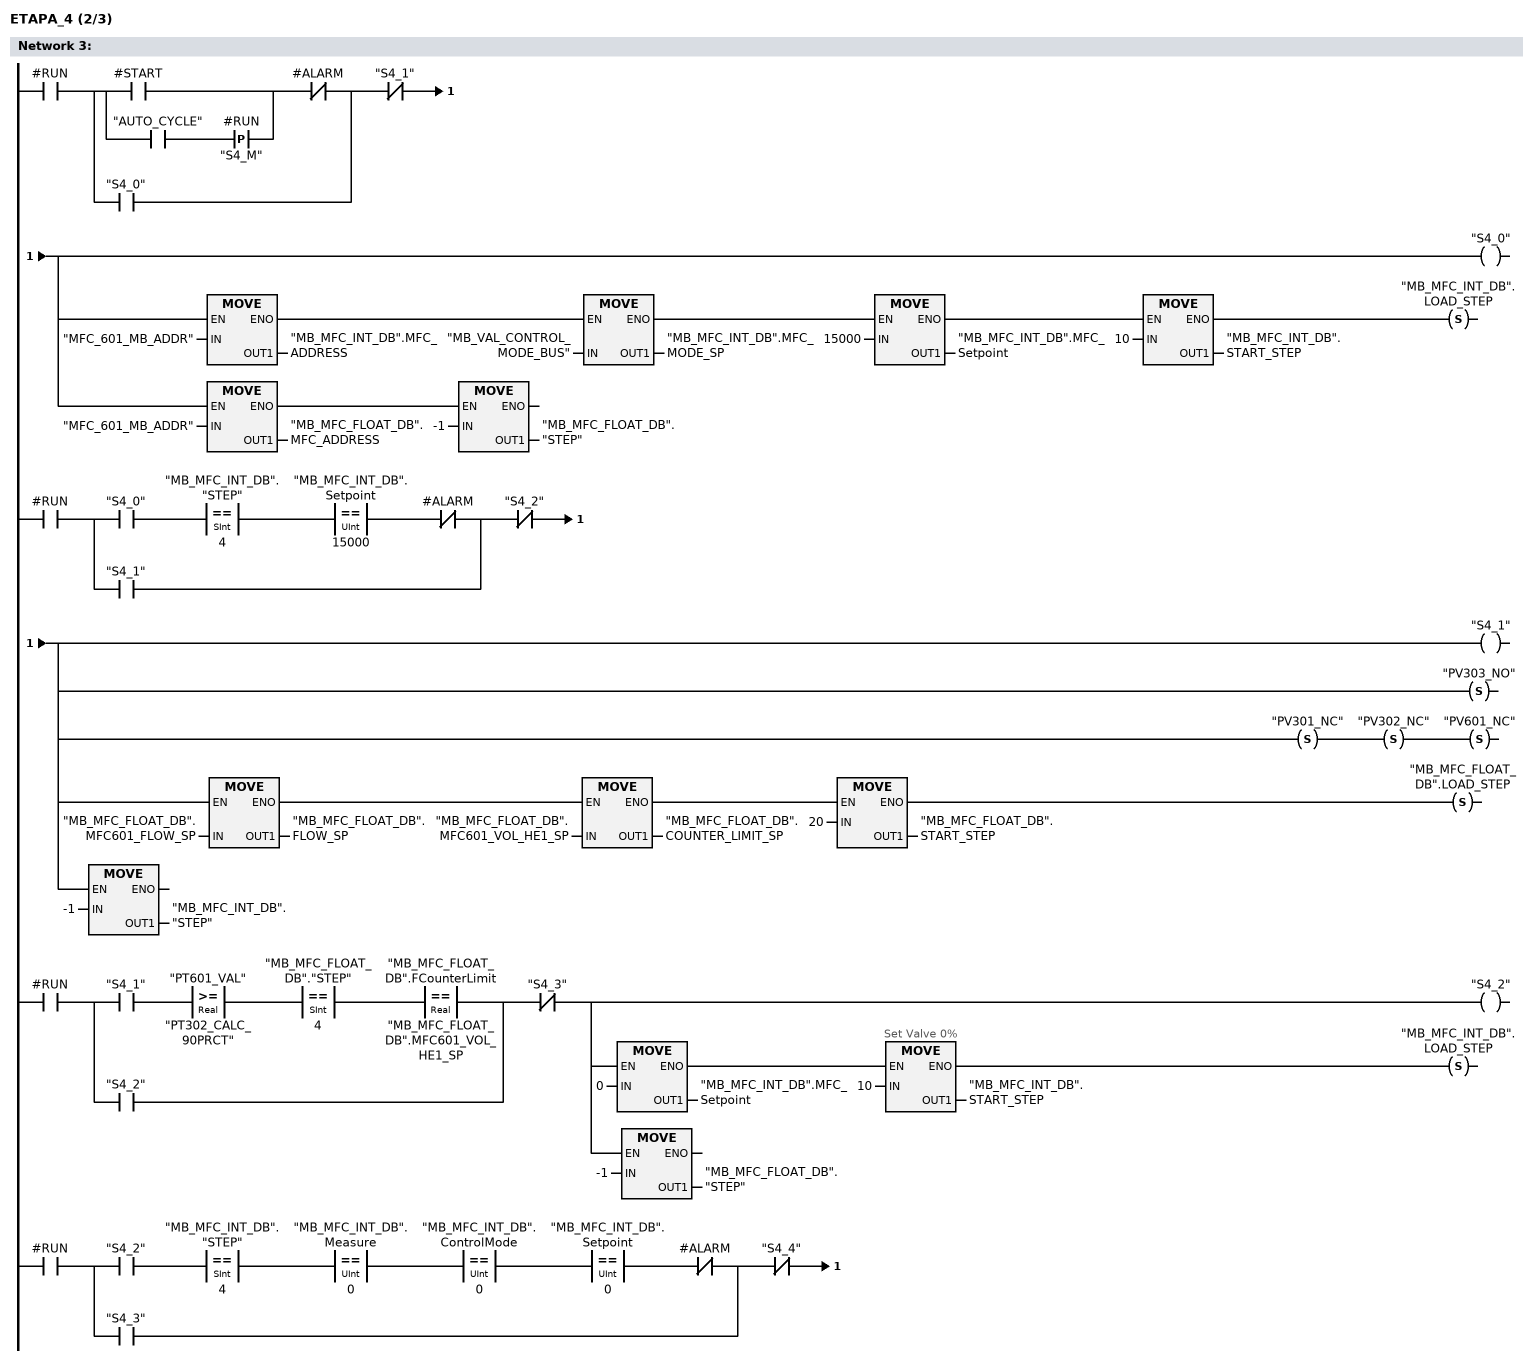
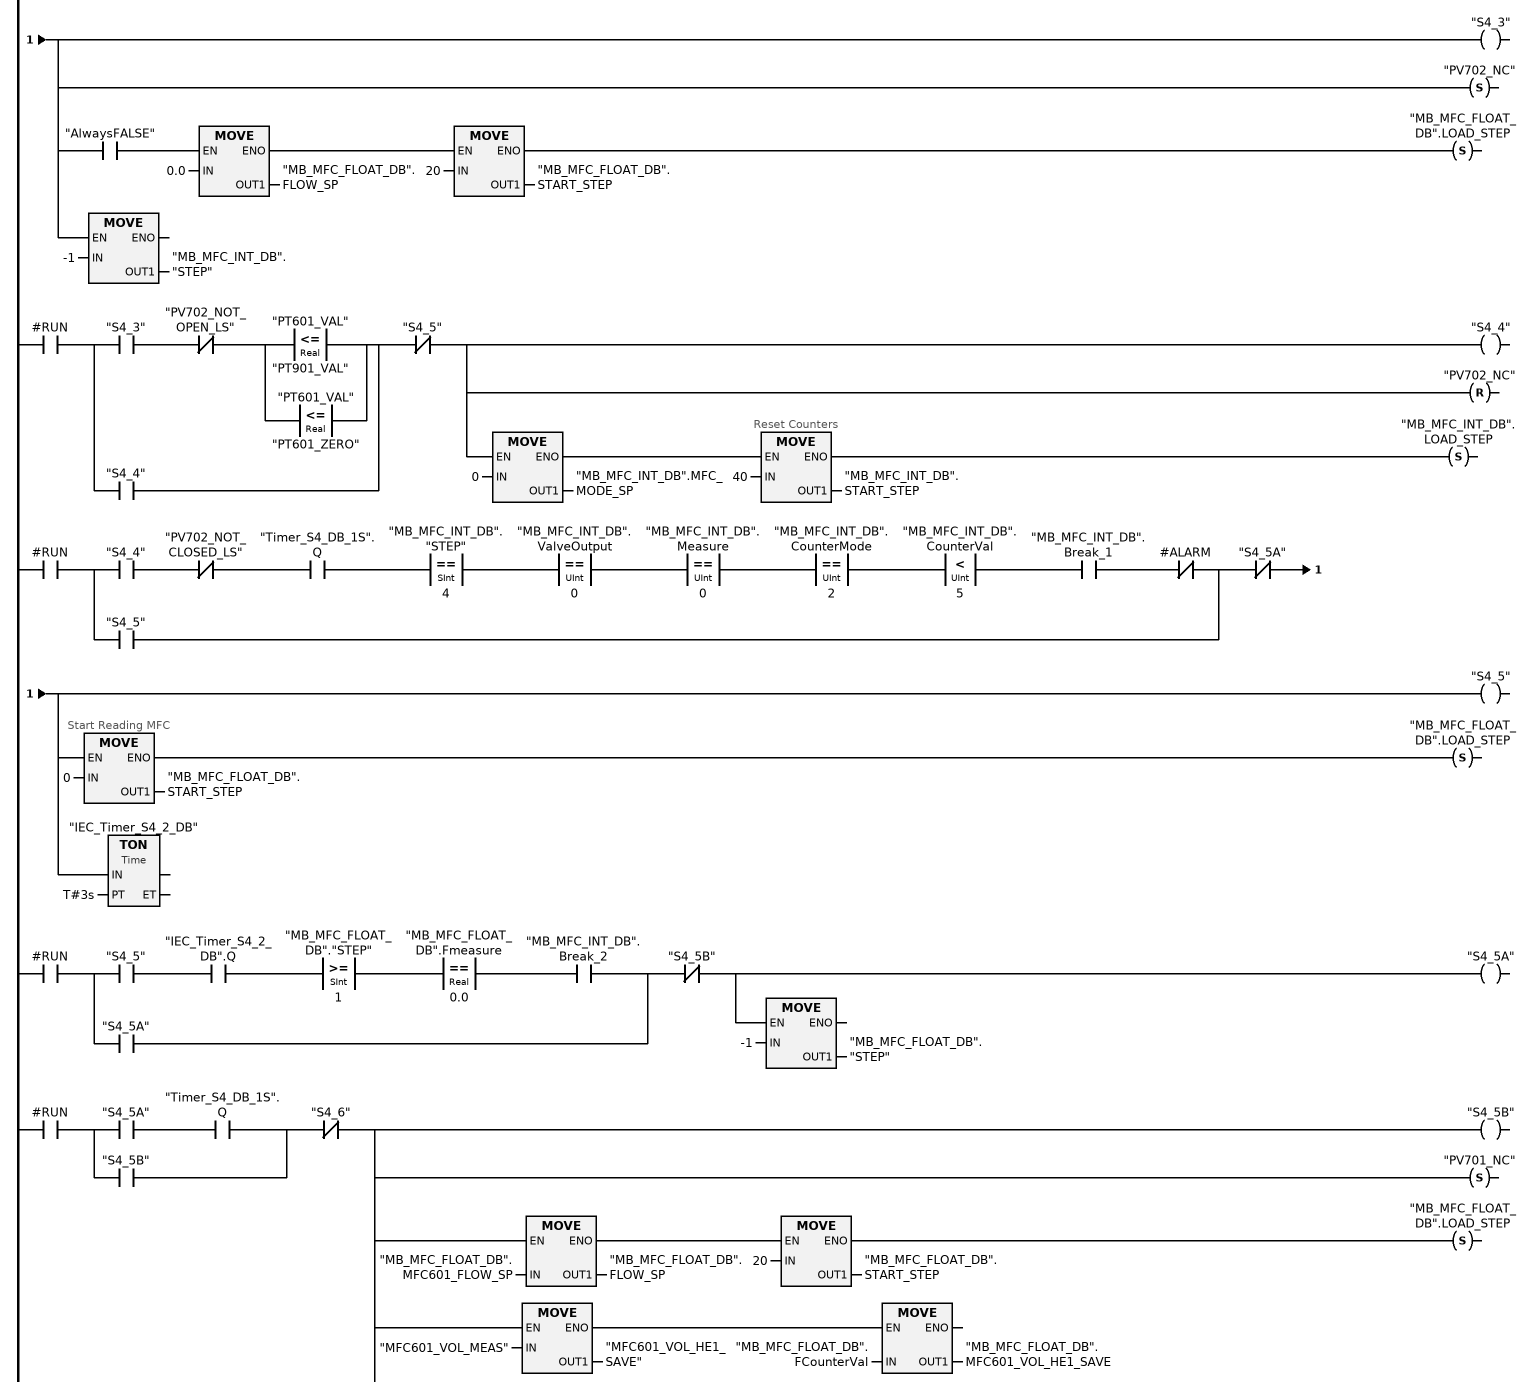
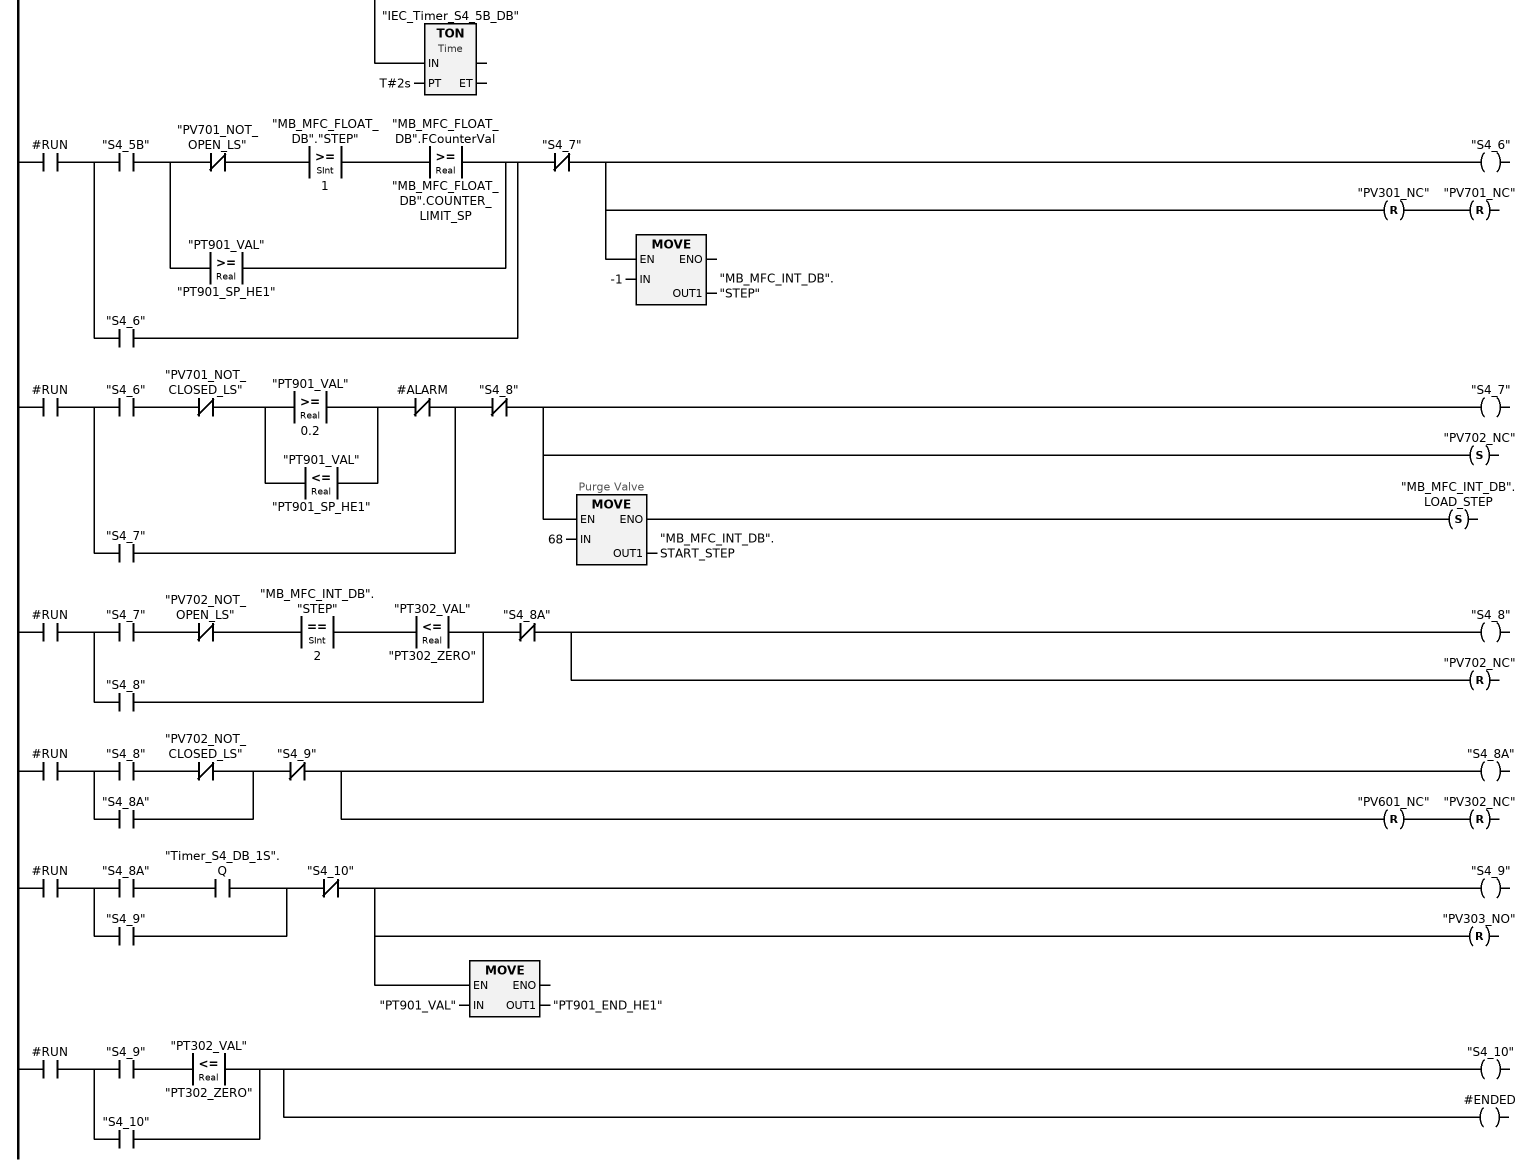
   #_w1 := #RUN AND "AUTO_CYCLE" AND #RUN AND NOT "S4_M";   // rising edge of #RUN
   "S4_M" := #RUN;
   "S4_0" := ((((#RUN AND #START) OR #_w1) AND NOT #ALARM) OR (#RUN AND "S4_0")) AND NOT "S4_1";
   IF "S4_0" THEN
       "MB_MFC_INT_DB".MFC_ADDRESS := "MFC_601_MB_ADDR";
       "MB_MFC_INT_DB".MFC_MODE_SP := "MB_VAL_CONTROL_MODE_BUS";
       "MB_MFC_INT_DB".MFC_Setpoint := 15000;
       "MB_MFC_INT_DB".START_STEP := 10;
       "MB_MFC_INT_DB".LOAD_STEP := TRUE;
       "MB_MFC_FLOAT_DB".MFC_ADDRESS := "MFC_601_MB_ADDR";
       "MB_MFC_FLOAT_DB"."STEP" := -1;
   END_IF;
   "S4_1" := #RUN AND (("S4_0" AND ("MB_MFC_INT_DB"."STEP" = 4) AND ("MB_MFC_INT_DB".Setpoint = 15000) AND NOT #ALARM) OR "S4_1") AND NOT "S4_2";
   IF "S4_1" THEN
       "PV303_NO" := TRUE;
       "PV301_NC" := TRUE;
       "PV302_NC" := TRUE;
       "PV601_NC" := TRUE;
       "MB_MFC_FLOAT_DB".FLOW_SP := "MB_MFC_FLOAT_DB".MFC601_FLOW_SP;
       "MB_MFC_FLOAT_DB".COUNTER_LIMIT_SP := "MB_MFC_FLOAT_DB".MFC601_VOL_HE1_SP;
       "MB_MFC_FLOAT_DB".START_STEP := 20;
       "MB_MFC_FLOAT_DB".LOAD_STEP := TRUE;
       "MB_MFC_INT_DB"."STEP" := -1;
   END_IF;
   "S4_2" := #RUN AND (("S4_1" AND ("PT601_VAL" >= "PT302_CALC_90PRCT") AND ("MB_MFC_FLOAT_DB"."STEP" = 4) AND ("MB_MFC_FLOAT_DB".FCounterLimit = "MB_MFC_FLOAT_DB".MFC601_VOL_HE1_SP)) OR "S4_2") AND NOT "S4_3";
   IF "S4_2" THEN
       "MB_MFC_INT_DB".MFC_Setpoint := 0;
       "MB_MFC_INT_DB".START_STEP := 10;   // Set Valve 0%
       "MB_MFC_INT_DB".LOAD_STEP := TRUE;
       "MB_MFC_FLOAT_DB"."STEP" := -1;
   END_IF;
   "S4_3" := #RUN AND (("S4_2" AND ("MB_MFC_INT_DB"."STEP" = 4) AND ("MB_MFC_INT_DB".Measure = 0) AND ("MB_MFC_INT_DB".ControlMode = 0) AND ("MB_MFC_INT_DB".Setpoint = 0) AND NOT #ALARM) OR "S4_3") AND NOT "S4_4";
   IF "S4_3" THEN "PV702_NC" := TRUE; END_IF;
   IF "S4_3" AND "AlwaysFALSE" THEN
       "MB_MFC_FLOAT_DB".FLOW_SP := 0.0;
       "MB_MFC_FLOAT_DB".START_STEP := 20;
       "MB_MFC_FLOAT_DB".LOAD_STEP := TRUE;
   END_IF;
   IF "S4_3" THEN "MB_MFC_INT_DB"."STEP" := -1; END_IF;
   "S4_4" := #RUN AND (("S4_3" AND NOT "PV702_NOT_OPEN_LS" AND (("PT601_VAL" <= "PT901_VAL") OR ("PT601_VAL" <= "PT601_ZERO"))) OR "S4_4") AND NOT "S4_5";
   IF "S4_4" THEN
       "PV702_NC" := FALSE;
       "MB_MFC_INT_DB".MFC_MODE_SP := 0;
       "MB_MFC_INT_DB".START_STEP := 40;   // Reset Counters
       "MB_MFC_INT_DB".LOAD_STEP := TRUE;
   END_IF;
   "S4_5" := #RUN AND (("S4_4" AND NOT "PV702_NOT_CLOSED_LS" AND "Timer_S4_DB_1S".Q AND ("MB_MFC_INT_DB"."STEP" = 4) AND ("MB_MFC_INT_DB".ValveOutput = 0) AND ("MB_MFC_INT_DB".Measure = 0) AND ("MB_MFC_INT_DB".CounterMode = 2) AND ("MB_MFC_INT_DB".CounterVal < 5) AND "MB_MFC_INT_DB".Break_1 AND NOT #ALARM) OR "S4_5") AND NOT "S4_5A";
   IF "S4_5" THEN
       "MB_MFC_FLOAT_DB".START_STEP := 0;   // Start Reading MFC
       "MB_MFC_FLOAT_DB".LOAD_STEP := TRUE;
   END_IF;
   "IEC_Timer_S4_2_DB".TON(IN := "S4_5", PT := T#3s);
   "S4_5A" := #RUN AND (("S4_5" AND "IEC_Timer_S4_2_DB".Q AND ("MB_MFC_FLOAT_DB"."STEP" >= 1) AND ("MB_MFC_FLOAT_DB".Fmeasure = 0.0) AND "MB_MFC_INT_DB".Break_2) OR "S4_5A") AND NOT "S4_5B";
   IF "S4_5A" THEN "MB_MFC_FLOAT_DB"."STEP" := -1; END_IF;
   "S4_5B" := #RUN AND (("S4_5A" AND "Timer_S4_DB_1S".Q) OR "S4_5B") AND NOT "S4_6";
   IF "S4_5B" THEN
       "PV701_NC" := TRUE;
       "MB_MFC_FLOAT_DB".FLOW_SP := "MB_MFC_FLOAT_DB".MFC601_FLOW_SP;
       "MB_MFC_FLOAT_DB".START_STEP := 20;
       "MB_MFC_FLOAT_DB".LOAD_STEP := TRUE;
       "MFC601_VOL_HE1_SAVE" := "MFC601_VOL_MEAS";
       "MB_MFC_FLOAT_DB".MFC601_VOL_HE1_SAVE := "MB_MFC_FLOAT_DB".FCounterVal;
   END_IF;
   "IEC_Timer_S4_5B_DB".TON(IN := "S4_5B", PT := T#2s);
   "S4_6" := #RUN AND (("S4_5B" AND ((NOT "PV701_NOT_OPEN_LS" AND ("MB_MFC_FLOAT_DB"."STEP" >= 1) AND ("MB_MFC_FLOAT_DB".FCounterVal >= "MB_MFC_FLOAT_DB".COUNTER_LIMIT_SP)) OR ("PT901_VAL" >= "PT901_SP_HE1"))) OR "S4_6") AND NOT "S4_7";
   IF "S4_6" THEN
       "PV301_NC" := FALSE;
       "PV701_NC" := FALSE;
       "MB_MFC_INT_DB"."STEP" := -1;
   END_IF;
   "S4_7" := #RUN AND (("S4_6" AND NOT "PV701_NOT_CLOSED_LS" AND (("PT901_VAL" >= 0.2) OR ("PT901_VAL" <= "PT901_SP_HE1")) AND NOT #ALARM) OR "S4_7") AND NOT "S4_8";
   IF "S4_7" THEN
       "PV702_NC" := TRUE;
       "MB_MFC_INT_DB".START_STEP := 68;   // Purge Valve
       "MB_MFC_INT_DB".LOAD_STEP := TRUE;
   END_IF;
   "S4_8" := #RUN AND (("S4_7" AND NOT "PV702_NOT_OPEN_LS" AND ("MB_MFC_INT_DB"."STEP" = 2) AND ("PT302_VAL" <= "PT302_ZERO")) OR "S4_8") AND NOT "S4_8A";
   IF "S4_8" THEN "PV702_NC" := FALSE; END_IF;
   "S4_8A" := #RUN AND (("S4_8" AND NOT "PV702_NOT_CLOSED_LS") OR "S4_8A") AND NOT "S4_9";
   IF "S4_8A" THEN
       "PV601_NC" := FALSE;
       "PV302_NC" := FALSE;
   END_IF;
   "S4_9" := #RUN AND (("S4_8A" AND "Timer_S4_DB_1S".Q) OR "S4_9") AND NOT "S4_10";
   IF "S4_9" THEN
       "PV303_NO" := FALSE;
       "PT901_END_HE1" := "PT901_VAL";
   END_IF;
   "S4_10" := #RUN AND (("S4_9" AND ("PT302_VAL" <= "PT302_ZERO")) OR "S4_10");
   #ENDED := "S4_10";
END_REGION

REGION Network 4
   // Timers
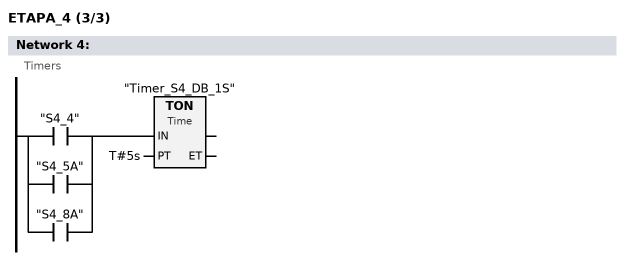
   "Timer_S4_DB_1S".TON(IN := "S4_4" OR "S4_5A" OR "S4_8A", PT := T#5s);
END_REGION
END_FUNCTION

FUNCTION "ETAPA_5" : Void   // FC6, LAD
{ S7_Optimized_Access := 'FALSE' }
VERSION : 0.1
// CICLO de INJECÇÃO - Varrimento Helio 2
   VAR_TEMP   // added for the SCL form of the ladder/FBD networks
      _w1 : Bool;
   END_VAR
BEGIN

REGION Network 1
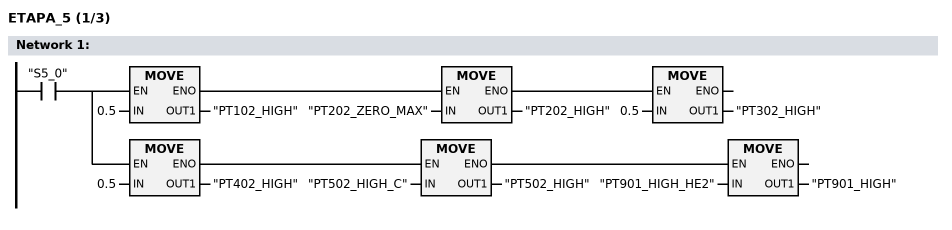
   RUNG wire#powerrail
      Contact( "S5_0" )
      wire#w1
      { S7_GenerateENO := "TRUE" } Move(in := 0.5, out1 => "PT102_HIGH")
      { S7_GenerateENO := "TRUE" } Move(in := "PT202_ZERO_MAX", out1 => "PT202_HIGH")
      { S7_GenerateENO := "TRUE" } Move(in := 0.5, out1 => "PT302_HIGH")
   END_RUNG
   RUNG wire#w1
      { S7_GenerateENO := "TRUE" } Move(in := 0.5, out1 => "PT402_HIGH")
      { S7_GenerateENO := "TRUE" } Move(in := "PT502_HIGH_C", out1 => "PT502_HIGH")
      { S7_GenerateENO := "TRUE" } Move(in := "PT901_HIGH_HE2", out1 => "PT901_HIGH")
   END_RUNG
   // the same network as SCL:
   // ENO of a box is taken as its EN; it also drops when the box reports an error
   IF "S5_0" THEN
       "PT102_HIGH" := 0.5;
       "PT202_HIGH" := "PT202_ZERO_MAX";
       "PT302_HIGH" := 0.5;
       "PT402_HIGH" := 0.5;
       "PT502_HIGH" := "PT502_HIGH_C";
       "PT901_HIGH" := "PT901_HIGH_HE2";
   END_IF;
END_REGION

REGION Network 2
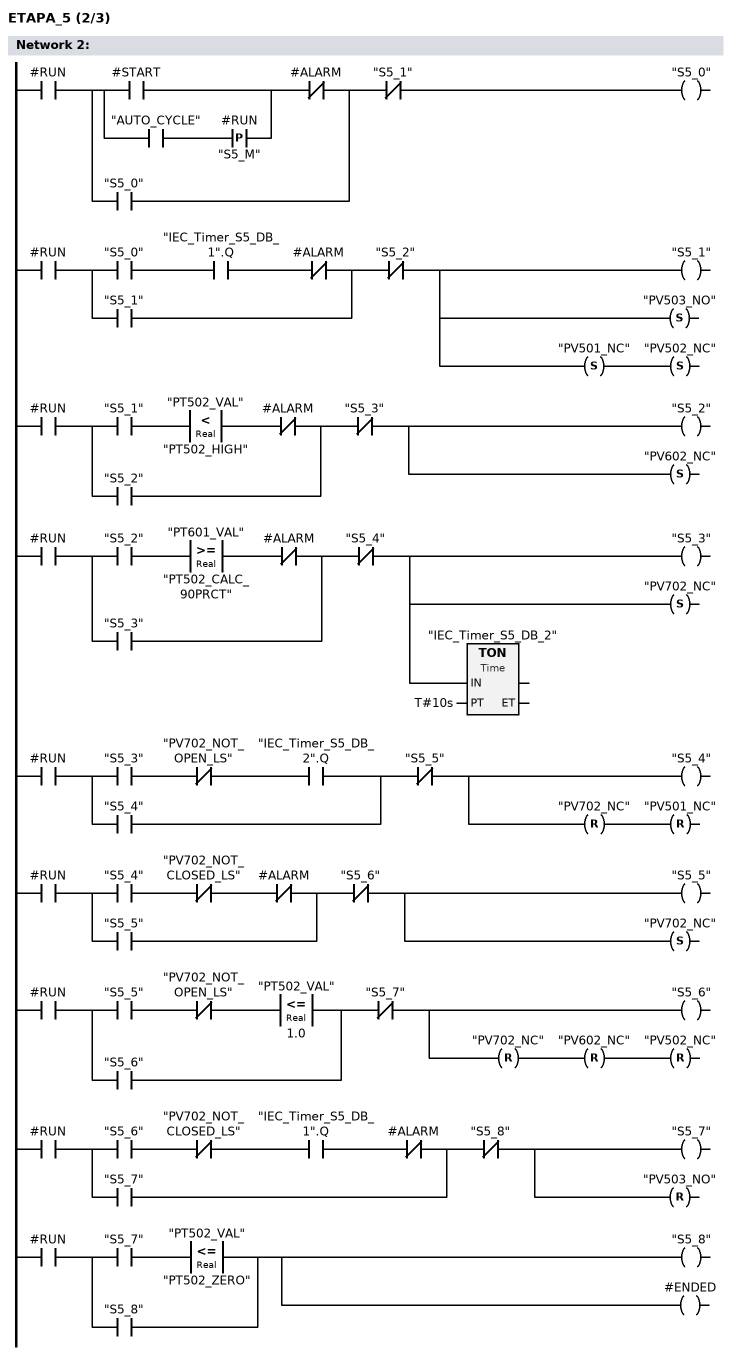
   #_w1 := #RUN AND "AUTO_CYCLE" AND #RUN AND NOT "S5_M";   // rising edge of #RUN
   "S5_M" := #RUN;
   "S5_0" := ((((#RUN AND #START) OR #_w1) AND NOT #ALARM) OR (#RUN AND "S5_0")) AND NOT "S5_1";
   "S5_1" := #RUN AND (("S5_0" AND "IEC_Timer_S5_DB_1".Q AND NOT #ALARM) OR "S5_1") AND NOT "S5_2";
   IF "S5_1" THEN
       "PV503_NO" := TRUE;
       "PV501_NC" := TRUE;
       "PV502_NC" := TRUE;
   END_IF;
   "S5_2" := #RUN AND (("S5_1" AND ("PT502_VAL" < "PT502_HIGH") AND NOT #ALARM) OR "S5_2") AND NOT "S5_3";
   IF "S5_2" THEN "PV602_NC" := TRUE; END_IF;
   "S5_3" := #RUN AND (("S5_2" AND ("PT601_VAL" >= "PT502_CALC_90PRCT") AND NOT #ALARM) OR "S5_3") AND NOT "S5_4";
   IF "S5_3" THEN "PV702_NC" := TRUE; END_IF;
   "IEC_Timer_S5_DB_2".TON(IN := "S5_3", PT := T#10s);
   "S5_4" := #RUN AND (("S5_3" AND NOT "PV702_NOT_OPEN_LS" AND "IEC_Timer_S5_DB_2".Q) OR "S5_4") AND NOT "S5_5";
   IF "S5_4" THEN
       "PV702_NC" := FALSE;
       "PV501_NC" := FALSE;
   END_IF;
   "S5_5" := #RUN AND (("S5_4" AND NOT "PV702_NOT_CLOSED_LS" AND NOT #ALARM) OR "S5_5") AND NOT "S5_6";
   IF "S5_5" THEN "PV702_NC" := TRUE; END_IF;
   "S5_6" := #RUN AND (("S5_5" AND NOT "PV702_NOT_OPEN_LS" AND ("PT502_VAL" <= 1.0)) OR "S5_6") AND NOT "S5_7";
   IF "S5_6" THEN
       "PV702_NC" := FALSE;
       "PV602_NC" := FALSE;
       "PV502_NC" := FALSE;
   END_IF;
   "S5_7" := #RUN AND (("S5_6" AND NOT "PV702_NOT_CLOSED_LS" AND "IEC_Timer_S5_DB_1".Q AND NOT #ALARM) OR "S5_7") AND NOT "S5_8";
   IF "S5_7" THEN "PV503_NO" := FALSE; END_IF;
   "S5_8" := #RUN AND (("S5_7" AND ("PT502_VAL" <= "PT502_ZERO")) OR "S5_8");
   #ENDED := "S5_8";
END_REGION

REGION Network 3
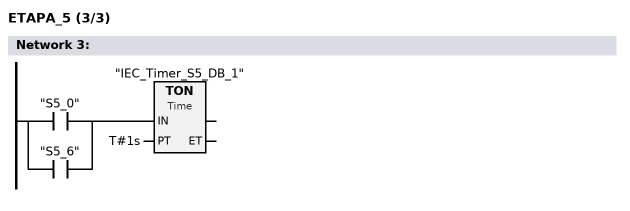
   "IEC_Timer_S5_DB_1".TON(IN := "S5_0" OR "S5_6", PT := T#1s);
END_REGION
END_FUNCTION

FUNCTION "ETAPA_6" : Void   // FC7, LAD
{ S7_Optimized_Access := 'FALSE' }
VERSION : 0.1
// CICLO de INJECÇÃO - injecção de Hidrogénio
   VAR_TEMP   // added for the SCL form of the ladder/FBD networks
      _w1 : Bool;
   END_VAR
BEGIN

REGION Network 1
   // Alarm PT Set Points
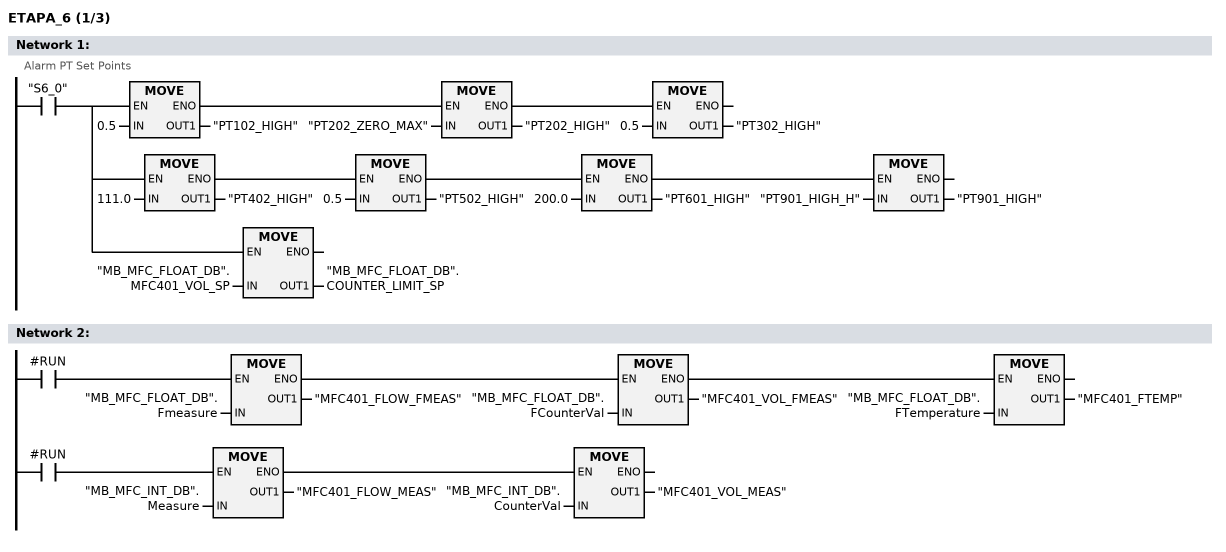
   RUNG wire#powerrail
      Contact( "S6_0" )
      wire#w1
      { S7_GenerateENO := "TRUE" } Move(in := 0.5, out1 => "PT102_HIGH")
      { S7_GenerateENO := "TRUE" } Move(in := "PT202_ZERO_MAX", out1 => "PT202_HIGH")
      { S7_GenerateENO := "TRUE" } Move(in := 0.5, out1 => "PT302_HIGH")
   END_RUNG
   RUNG wire#w1
      { S7_GenerateENO := "TRUE" } Move(in := 111.0, out1 => "PT402_HIGH")
      { S7_GenerateENO := "TRUE" } Move(in := 0.5, out1 => "PT502_HIGH")
      { S7_GenerateENO := "TRUE" } Move(in := 200.0, out1 => "PT601_HIGH")
      { S7_GenerateENO := "TRUE" } Move(in := "PT901_HIGH_H", out1 => "PT901_HIGH")
   END_RUNG
   RUNG wire#w1
      Move(in := "MB_MFC_FLOAT_DB".MFC401_VOL_SP, out1 => "MB_MFC_FLOAT_DB".COUNTER_LIMIT_SP)
   END_RUNG
   // the same network as SCL:
   // ENO of a box is taken as its EN; it also drops when the box reports an error
   IF "S6_0" THEN
       "PT102_HIGH" := 0.5;
       "PT202_HIGH" := "PT202_ZERO_MAX";
       "PT302_HIGH" := 0.5;
       "PT402_HIGH" := 111.0;
       "PT502_HIGH" := 0.5;
       "PT601_HIGH" := 200.0;
       "PT901_HIGH" := "PT901_HIGH_H";
       "MB_MFC_FLOAT_DB".COUNTER_LIMIT_SP := "MB_MFC_FLOAT_DB".MFC401_VOL_SP;
   END_IF;
END_REGION

REGION Network 2
   RUNG wire#powerrail
      Contact( #RUN )
      { S7_GenerateENO := "TRUE" } Move(in := "MB_MFC_FLOAT_DB".Fmeasure, out1 => "MFC401_FLOW_FMEAS")
      { S7_GenerateENO := "TRUE" } Move(in := "MB_MFC_FLOAT_DB".FCounterVal, out1 => "MFC401_VOL_FMEAS")
      { S7_GenerateENO := "TRUE" } Move(in := "MB_MFC_FLOAT_DB".FTemperature, out1 => "MFC401_FTEMP")
   END_RUNG
   RUNG wire#powerrail
      Contact( #RUN )
      { S7_GenerateENO := "TRUE" } Move(in := "MB_MFC_INT_DB".Measure, out1 => "MFC401_FLOW_MEAS")
      { S7_GenerateENO := "TRUE" } Move(in := "MB_MFC_INT_DB".CounterVal, out1 => "MFC401_VOL_MEAS")
   END_RUNG
   // the same network as SCL:
   // ENO of a box is taken as its EN; it also drops when the box reports an error
   IF #RUN THEN
       "MFC401_FLOW_FMEAS" := "MB_MFC_FLOAT_DB".Fmeasure;
       "MFC401_VOL_FMEAS" := "MB_MFC_FLOAT_DB".FCounterVal;
       "MFC401_FTEMP" := "MB_MFC_FLOAT_DB".FTemperature;
       "MFC401_FLOW_MEAS" := "MB_MFC_INT_DB".Measure;
       "MFC401_VOL_MEAS" := "MB_MFC_INT_DB".CounterVal;
   END_IF;
END_REGION

REGION Network 3
   // Logica do ciclo 6
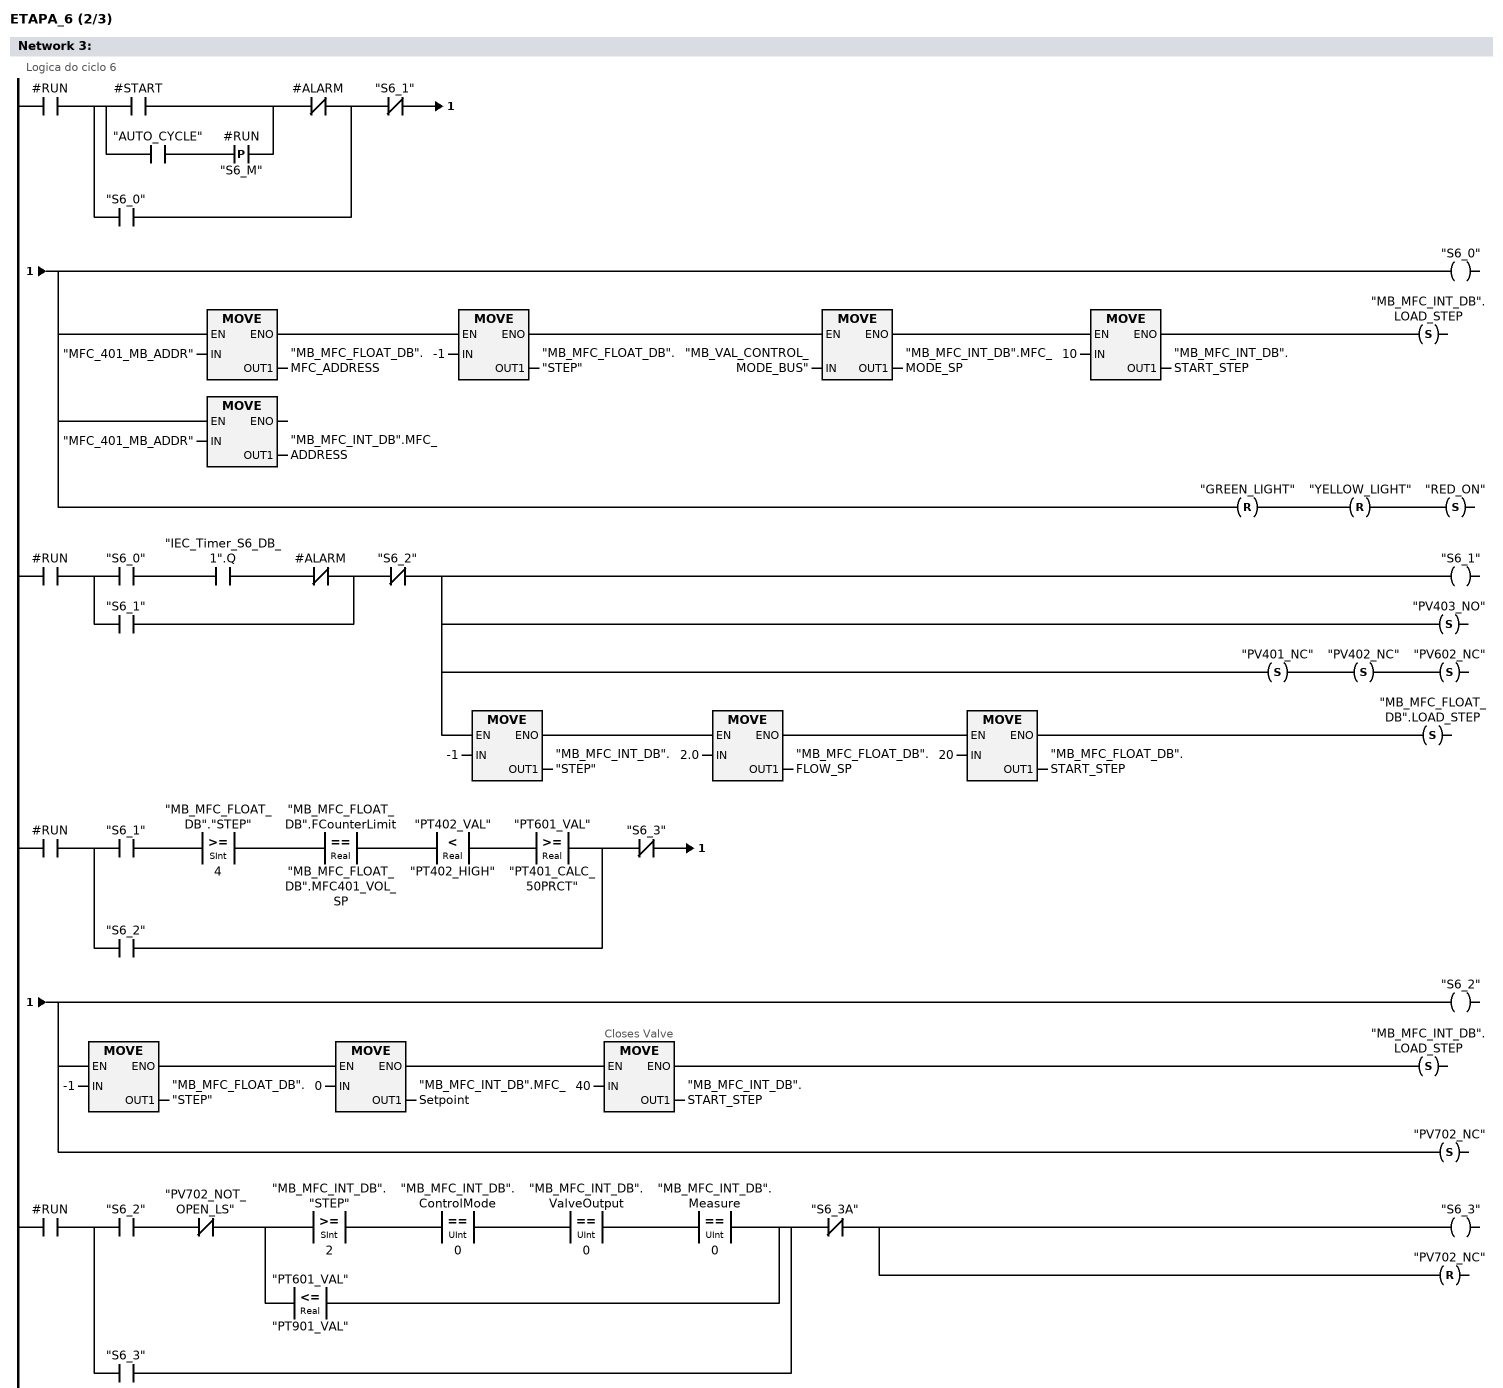
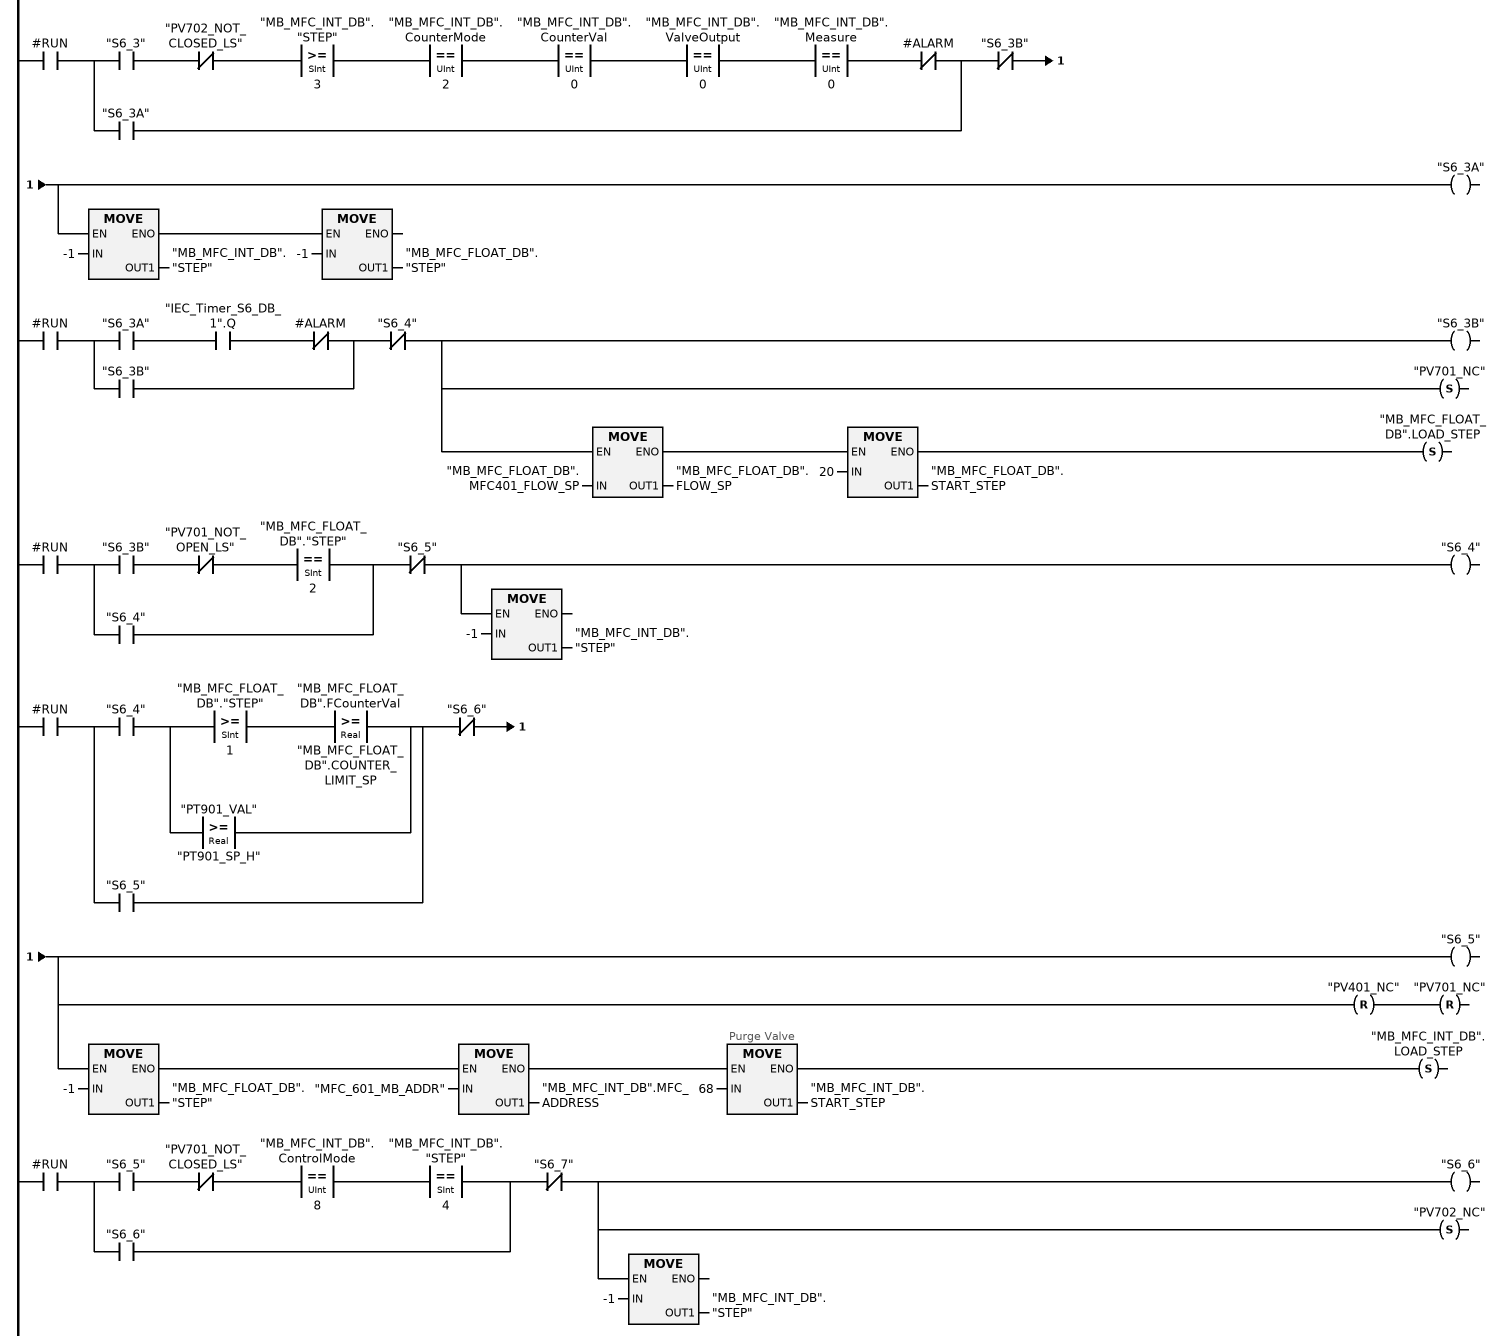
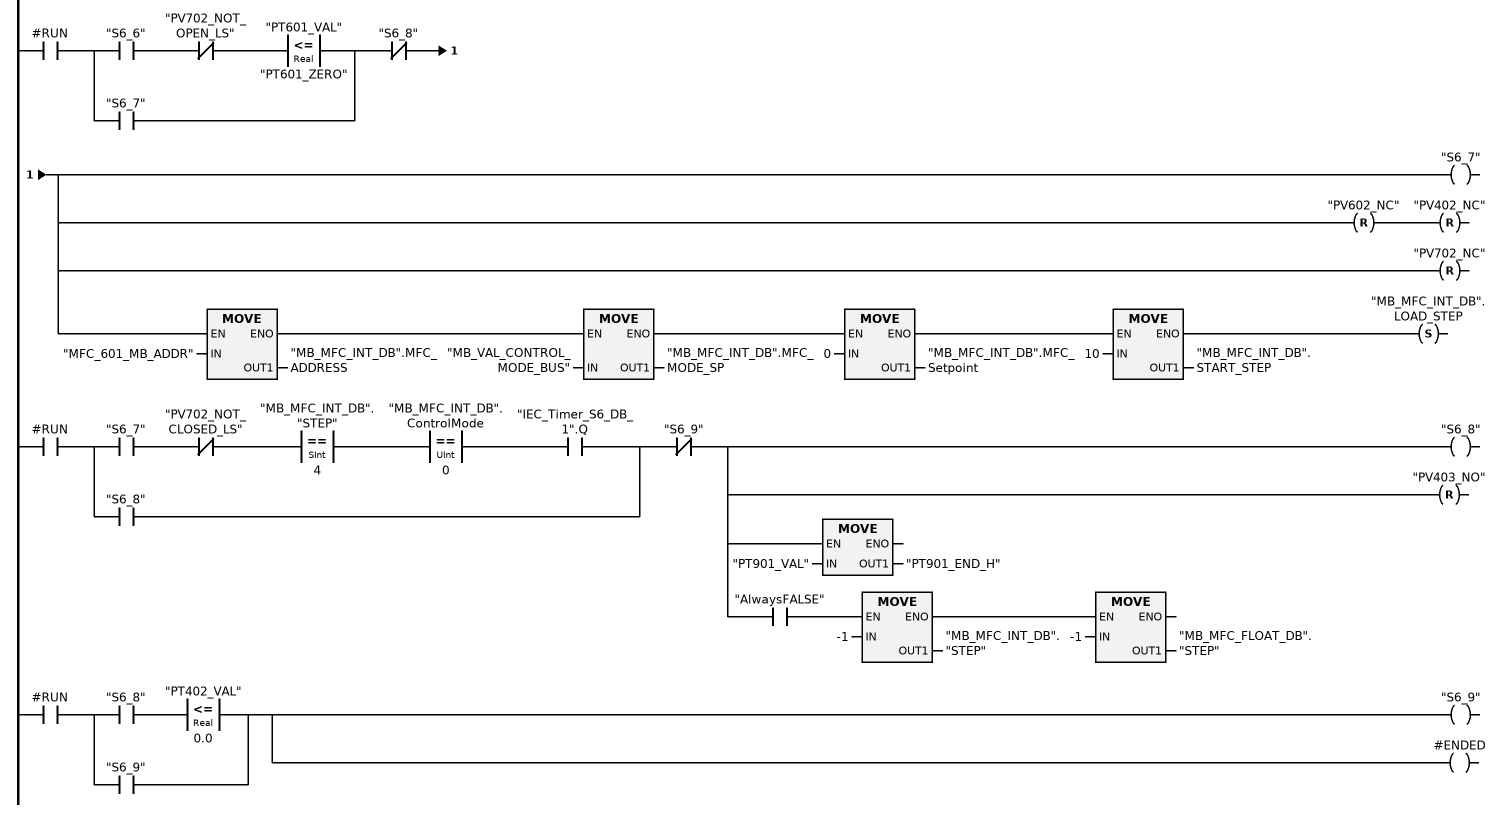
   RUNG wire#powerrail
      Contact( #RUN )
      wire#w1
      Contact( #START )
      wire#w2
      I_Contact( #ALARM )
      wire#w3
      I_Contact( "S6_1" )
      wire#w4
      Coil( "S6_0" )
   END_RUNG
   RUNG wire#w1
      Contact( "AUTO_CYCLE" )
      P_Contact(operand := #RUN, bit := "S6_M")
   END_RUNG wire#w2
   RUNG wire#w1
      Contact( "S6_0" )
   END_RUNG wire#w3
   RUNG wire#w4
      Move(in := "MFC_401_MB_ADDR", out1 => "MB_MFC_FLOAT_DB".MFC_ADDRESS)
      Move(in := -1, out1 => "MB_MFC_FLOAT_DB"."STEP")
      Move(in := "MB_VAL_CONTROL_MODE_BUS", out1 => "MB_MFC_INT_DB".MFC_MODE_SP)
      Move(in := 10, out1 => "MB_MFC_INT_DB".START_STEP)
      S_Coil( "MB_MFC_INT_DB".LOAD_STEP )
   END_RUNG
   RUNG wire#w4
      Move(in := "MFC_401_MB_ADDR", out1 => "MB_MFC_INT_DB".MFC_ADDRESS)
   END_RUNG
   RUNG wire#w4
      R_Coil( "GREEN_LIGHT" )
      R_Coil( "YELLOW_LIGHT" )
      S_Coil( "RED_ON" )
   END_RUNG
   RUNG wire#powerrail
      Contact( #RUN )
      wire#w5
      Contact( "S6_0" )
      Contact( "IEC_Timer_S6_DB_1".Q )
      I_Contact( #ALARM )
      wire#w6
      I_Contact( "S6_2" )
      wire#w7
      Coil( "S6_1" )
   END_RUNG
   RUNG wire#w5
      Contact( "S6_1" )
   END_RUNG wire#w6
   RUNG wire#w7
      S_Coil( "PV403_NO" )
   END_RUNG
   RUNG wire#w7
      S_Coil( "PV401_NC" )
      S_Coil( "PV402_NC" )
      S_Coil( "PV602_NC" )
   END_RUNG
   RUNG wire#w7
      Move(in := -1, out1 => "MB_MFC_INT_DB"."STEP")
      Move(in := 2.0, out1 => "MB_MFC_FLOAT_DB".FLOW_SP)
      Move(in := 20, out1 => "MB_MFC_FLOAT_DB".START_STEP)
      S_Coil( "MB_MFC_FLOAT_DB".LOAD_STEP )
   END_RUNG
   RUNG wire#powerrail
      Contact( #RUN )
      wire#w8
      Contact( "S6_1" )
      { S7_Templates := "SrcType := SInt" } GE_Contact(in1 := "MB_MFC_FLOAT_DB"."STEP", in2 := 4)